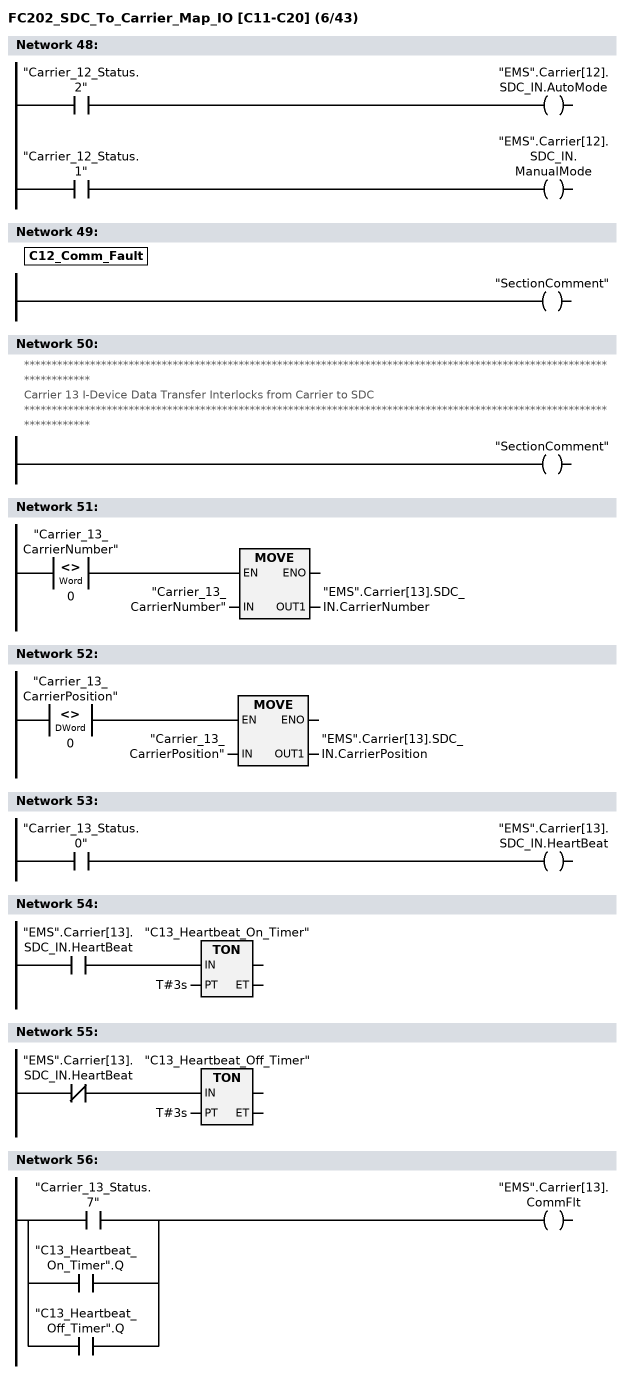
   RUNG wire#powerrail
      Contact( "Carrier_12_Status.2" )
      Coil( "EMS".Carrier[12].SDC_IN.AutoMode )
   END_RUNG
   RUNG wire#powerrail
      Contact( "Carrier_12_Status.1" )
      Coil( "EMS".Carrier[12].SDC_IN.ManualMode )
   END_RUNG
   // the same network as SCL:
   "EMS".Carrier[12].SDC_IN.AutoMode := "Carrier_12_Status.2";
   "EMS".Carrier[12].SDC_IN.ManualMode := "Carrier_12_Status.1";
END_REGION

REGION Network 49
   Label( C12_Comm_Fault )
   RUNG wire#powerrail
      Coil( "SectionComment" )
   END_RUNG
   // the same network as SCL:
   C12_Comm_Fault:
   "SectionComment" := TRUE;
END_REGION

REGION Network 50
   // **********************************************************************************************************************
   // 
   // Carrier 13 I-Device Data Transfer Interlocks from Carrier to SDC
   // 
   // **********************************************************************************************************************
   RUNG wire#powerrail
      Coil( "SectionComment" )
   END_RUNG
   // the same network as SCL:
   "SectionComment" := TRUE;
END_REGION

REGION Network 51
   RUNG wire#powerrail
      { S7_Templates := "SrcType := Word" } NE_Contact(in1 := "Carrier_13_CarrierNumber", in2 := 0)
      Move(in := "Carrier_13_CarrierNumber", out1 => "EMS".Carrier[13].SDC_IN.CarrierNumber)
   END_RUNG
   // the same network as SCL:
   IF "Carrier_13_CarrierNumber" <> 0 THEN
       "EMS".Carrier[13].SDC_IN.CarrierNumber := "Carrier_13_CarrierNumber";
   END_IF;
END_REGION

REGION Network 52
   RUNG wire#powerrail
      { S7_Templates := "SrcType := DWord" } NE_Contact(in1 := "Carrier_13_CarrierPosition", in2 := 0)
      Move(in := "Carrier_13_CarrierPosition", out1 => "EMS".Carrier[13].SDC_IN.CarrierPosition)
   END_RUNG
   // the same network as SCL:
   IF "Carrier_13_CarrierPosition" <> 0 THEN
       "EMS".Carrier[13].SDC_IN.CarrierPosition := "Carrier_13_CarrierPosition";
   END_IF;
END_REGION

REGION Network 53
   RUNG wire#powerrail
      Contact( "Carrier_13_Status.0" )
      Coil( "EMS".Carrier[13].SDC_IN.HeartBeat )
   END_RUNG
   // the same network as SCL:
   "EMS".Carrier[13].SDC_IN.HeartBeat := "Carrier_13_Status.0";
END_REGION

REGION Network 54
   "C13_Heartbeat_On_Timer".TON(IN := "EMS".Carrier[13].SDC_IN.HeartBeat, PT := T#3s);
END_REGION

REGION Network 55
   "C13_Heartbeat_Off_Timer".TON(IN := NOT "EMS".Carrier[13].SDC_IN.HeartBeat, PT := T#3s);
END_REGION

REGION Network 56
   RUNG wire#powerrail
      Contact( "Carrier_13_Status.7" )
      wire#w1
      Coil( "EMS".Carrier[13].CommFlt )
   END_RUNG
   RUNG wire#powerrail
      Contact( "C13_Heartbeat_On_Timer".Q )
   END_RUNG wire#w1
   RUNG wire#powerrail
      Contact( "C13_Heartbeat_Off_Timer".Q )
   END_RUNG wire#w1
   // the same network as SCL:
   "EMS".Carrier[13].CommFlt := "Carrier_13_Status.7" OR "C13_Heartbeat_On_Timer".Q OR "C13_Heartbeat_Off_Timer".Q;
END_REGION

REGION Network 57
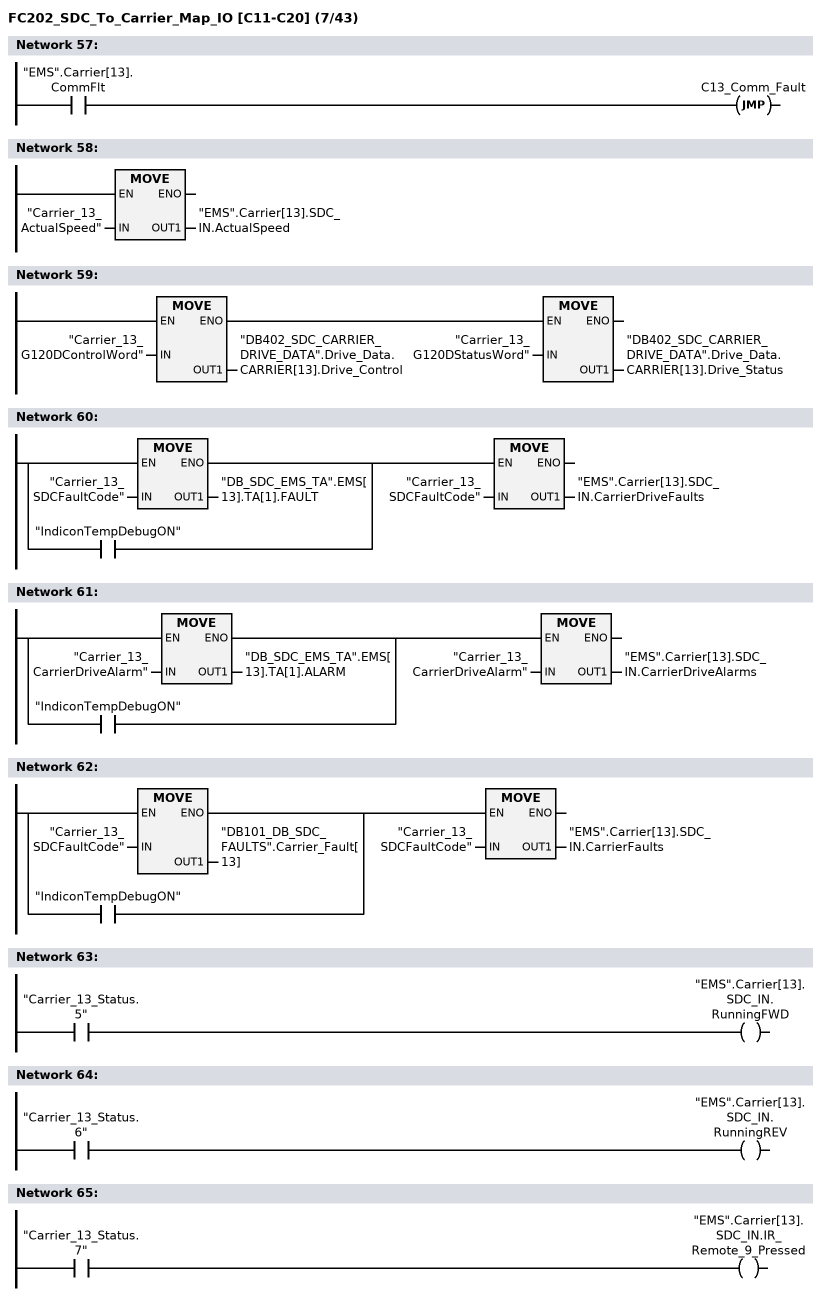
   RUNG wire#powerrail
      Contact( "EMS".Carrier[13].CommFlt )
      JumpCoil( C13_Comm_Fault )
   END_RUNG
   // the same network as SCL:
   IF "EMS".Carrier[13].CommFlt THEN GOTO C13_Comm_Fault; END_IF;
END_REGION

REGION Network 58
   RUNG wire#powerrail
      Move(in := "Carrier_13_ActualSpeed", out1 => "EMS".Carrier[13].SDC_IN.ActualSpeed)
   END_RUNG
   // the same network as SCL:
   "EMS".Carrier[13].SDC_IN.ActualSpeed := "Carrier_13_ActualSpeed";
END_REGION

REGION Network 59
   RUNG wire#powerrail
      Move(in := "Carrier_13_G120DControlWord", out1 => "DB402_SDC_CARRIER_DRIVE_DATA".Drive_Data.CARRIER[13].Drive_Control)
      Move(in := "Carrier_13_G120DStatusWord", out1 => "DB402_SDC_CARRIER_DRIVE_DATA".Drive_Data.CARRIER[13].Drive_Status)
   END_RUNG
   // the same network as SCL:
   "DB402_SDC_CARRIER_DRIVE_DATA".Drive_Data.CARRIER[13].Drive_Control := "Carrier_13_G120DControlWord";
   "DB402_SDC_CARRIER_DRIVE_DATA".Drive_Data.CARRIER[13].Drive_Status := "Carrier_13_G120DStatusWord";
END_REGION

REGION Network 60
   RUNG wire#powerrail
      Move(in := "Carrier_13_SDCFaultCode", out1 => "DB_SDC_EMS_TA".EMS[13].TA[1].FAULT)
      wire#w1
      Move(in := "Carrier_13_SDCFaultCode", out1 => "EMS".Carrier[13].SDC_IN.CarrierDriveFaults)
   END_RUNG
   RUNG wire#powerrail
      Contact( "IndiconTempDebugON" )
   END_RUNG wire#w1
   // the same network as SCL:
   "DB_SDC_EMS_TA".EMS[13].TA[1].FAULT := "Carrier_13_SDCFaultCode";
   IF TRUE OR "IndiconTempDebugON" THEN
       "EMS".Carrier[13].SDC_IN.CarrierDriveFaults := "Carrier_13_SDCFaultCode";
   END_IF;
END_REGION

REGION Network 61
   RUNG wire#powerrail
      Move(in := "Carrier_13_CarrierDriveAlarm", out1 => "DB_SDC_EMS_TA".EMS[13].TA[1].ALARM)
      wire#w1
      Move(in := "Carrier_13_CarrierDriveAlarm", out1 => "EMS".Carrier[13].SDC_IN.CarrierDriveAlarms)
   END_RUNG
   RUNG wire#powerrail
      Contact( "IndiconTempDebugON" )
   END_RUNG wire#w1
   // the same network as SCL:
   "DB_SDC_EMS_TA".EMS[13].TA[1].ALARM := "Carrier_13_CarrierDriveAlarm";
   IF TRUE OR "IndiconTempDebugON" THEN
       "EMS".Carrier[13].SDC_IN.CarrierDriveAlarms := "Carrier_13_CarrierDriveAlarm";
   END_IF;
END_REGION

REGION Network 62
   RUNG wire#powerrail
      Move(in := "Carrier_13_SDCFaultCode", out1 => "DB101_DB_SDC_FAULTS".Carrier_Fault[13])
      wire#w1
      Move(in := "Carrier_13_SDCFaultCode", out1 => "EMS".Carrier[13].SDC_IN.CarrierFaults)
   END_RUNG
   RUNG wire#powerrail
      Contact( "IndiconTempDebugON" )
   END_RUNG wire#w1
   // the same network as SCL:
   "DB101_DB_SDC_FAULTS".Carrier_Fault[13] := "Carrier_13_SDCFaultCode";
   IF TRUE OR "IndiconTempDebugON" THEN
       "EMS".Carrier[13].SDC_IN.CarrierFaults := "Carrier_13_SDCFaultCode";
   END_IF;
END_REGION

REGION Network 63
   RUNG wire#powerrail
      Contact( "Carrier_13_Status.5" )
      Coil( "EMS".Carrier[13].SDC_IN.RunningFWD )
   END_RUNG
   // the same network as SCL:
   "EMS".Carrier[13].SDC_IN.RunningFWD := "Carrier_13_Status.5";
END_REGION

REGION Network 64
   RUNG wire#powerrail
      Contact( "Carrier_13_Status.6" )
      Coil( "EMS".Carrier[13].SDC_IN.RunningREV )
   END_RUNG
   // the same network as SCL:
   "EMS".Carrier[13].SDC_IN.RunningREV := "Carrier_13_Status.6";
END_REGION

REGION Network 65
   RUNG wire#powerrail
      Contact( "Carrier_13_Status.7" )
      Coil( "EMS".Carrier[13].SDC_IN.IR_Remote_9_Pressed )
   END_RUNG
   // the same network as SCL:
   "EMS".Carrier[13].SDC_IN.IR_Remote_9_Pressed := "Carrier_13_Status.7";
END_REGION

REGION Network 66
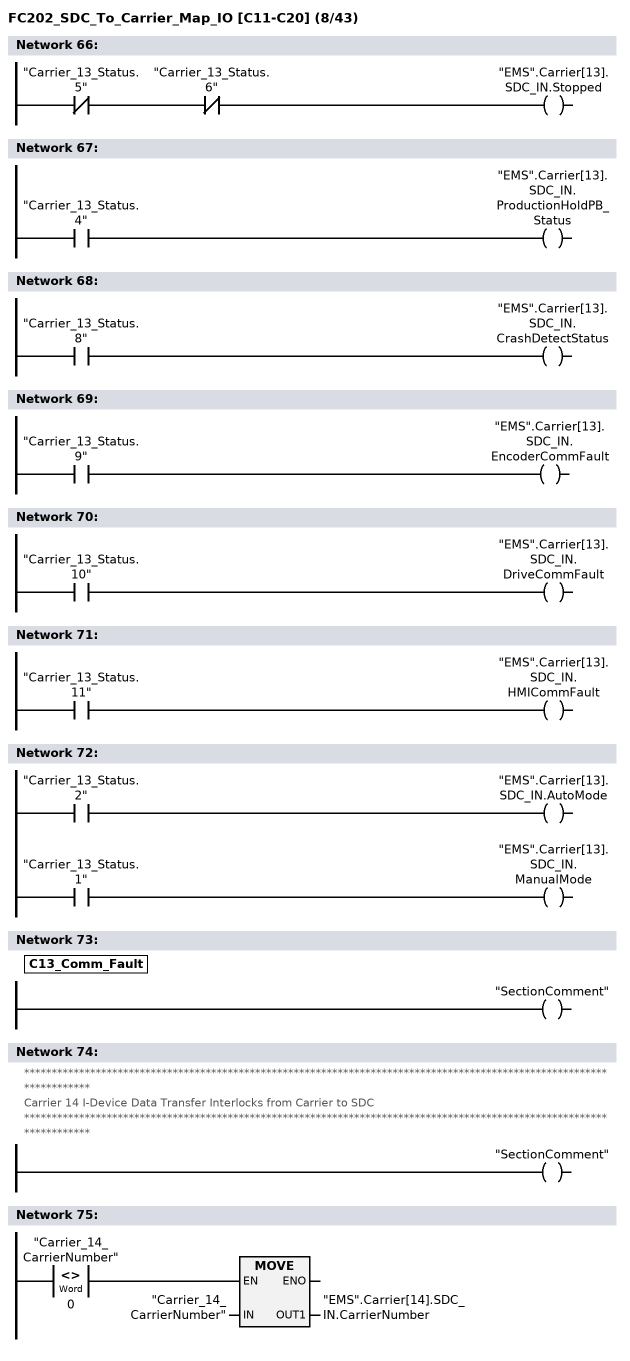
   RUNG wire#powerrail
      I_Contact( "Carrier_13_Status.5" )
      I_Contact( "Carrier_13_Status.6" )
      Coil( "EMS".Carrier[13].SDC_IN.Stopped )
   END_RUNG
   // the same network as SCL:
   "EMS".Carrier[13].SDC_IN.Stopped := NOT "Carrier_13_Status.5" AND NOT "Carrier_13_Status.6";
END_REGION

REGION Network 67
   RUNG wire#powerrail
      Contact( "Carrier_13_Status.4" )
      Coil( "EMS".Carrier[13].SDC_IN.ProductionHoldPB_Status )
   END_RUNG
   // the same network as SCL:
   "EMS".Carrier[13].SDC_IN.ProductionHoldPB_Status := "Carrier_13_Status.4";
END_REGION

REGION Network 68
   RUNG wire#powerrail
      Contact( "Carrier_13_Status.8" )
      Coil( "EMS".Carrier[13].SDC_IN.CrashDetectStatus )
   END_RUNG
   // the same network as SCL:
   "EMS".Carrier[13].SDC_IN.CrashDetectStatus := "Carrier_13_Status.8";
END_REGION

REGION Network 69
   RUNG wire#powerrail
      Contact( "Carrier_13_Status.9" )
      Coil( "EMS".Carrier[13].SDC_IN.EncoderCommFault )
   END_RUNG
   // the same network as SCL:
   "EMS".Carrier[13].SDC_IN.EncoderCommFault := "Carrier_13_Status.9";
END_REGION

REGION Network 70
   RUNG wire#powerrail
      Contact( "Carrier_13_Status.10" )
      Coil( "EMS".Carrier[13].SDC_IN.DriveCommFault )
   END_RUNG
   // the same network as SCL:
   "EMS".Carrier[13].SDC_IN.DriveCommFault := "Carrier_13_Status.10";
END_REGION

REGION Network 71
   RUNG wire#powerrail
      Contact( "Carrier_13_Status.11" )
      Coil( "EMS".Carrier[13].SDC_IN.HMICommFault )
   END_RUNG
   // the same network as SCL:
   "EMS".Carrier[13].SDC_IN.HMICommFault := "Carrier_13_Status.11";
END_REGION

REGION Network 72
   RUNG wire#powerrail
      Contact( "Carrier_13_Status.2" )
      Coil( "EMS".Carrier[13].SDC_IN.AutoMode )
   END_RUNG
   RUNG wire#powerrail
      Contact( "Carrier_13_Status.1" )
      Coil( "EMS".Carrier[13].SDC_IN.ManualMode )
   END_RUNG
   // the same network as SCL:
   "EMS".Carrier[13].SDC_IN.AutoMode := "Carrier_13_Status.2";
   "EMS".Carrier[13].SDC_IN.ManualMode := "Carrier_13_Status.1";
END_REGION

REGION Network 73
   Label( C13_Comm_Fault )
   RUNG wire#powerrail
      Coil( "SectionComment" )
   END_RUNG
   // the same network as SCL:
   C13_Comm_Fault:
   "SectionComment" := TRUE;
END_REGION

REGION Network 74
   // **********************************************************************************************************************
   // 
   // Carrier 14 I-Device Data Transfer Interlocks from Carrier to SDC
   // 
   // **********************************************************************************************************************
   RUNG wire#powerrail
      Coil( "SectionComment" )
   END_RUNG
   // the same network as SCL:
   "SectionComment" := TRUE;
END_REGION

REGION Network 75
   RUNG wire#powerrail
      { S7_Templates := "SrcType := Word" } NE_Contact(in1 := "Carrier_14_CarrierNumber", in2 := 0)
      Move(in := "Carrier_14_CarrierNumber", out1 => "EMS".Carrier[14].SDC_IN.CarrierNumber)
   END_RUNG
   // the same network as SCL:
   IF "Carrier_14_CarrierNumber" <> 0 THEN
       "EMS".Carrier[14].SDC_IN.CarrierNumber := "Carrier_14_CarrierNumber";
   END_IF;
END_REGION

REGION Network 76
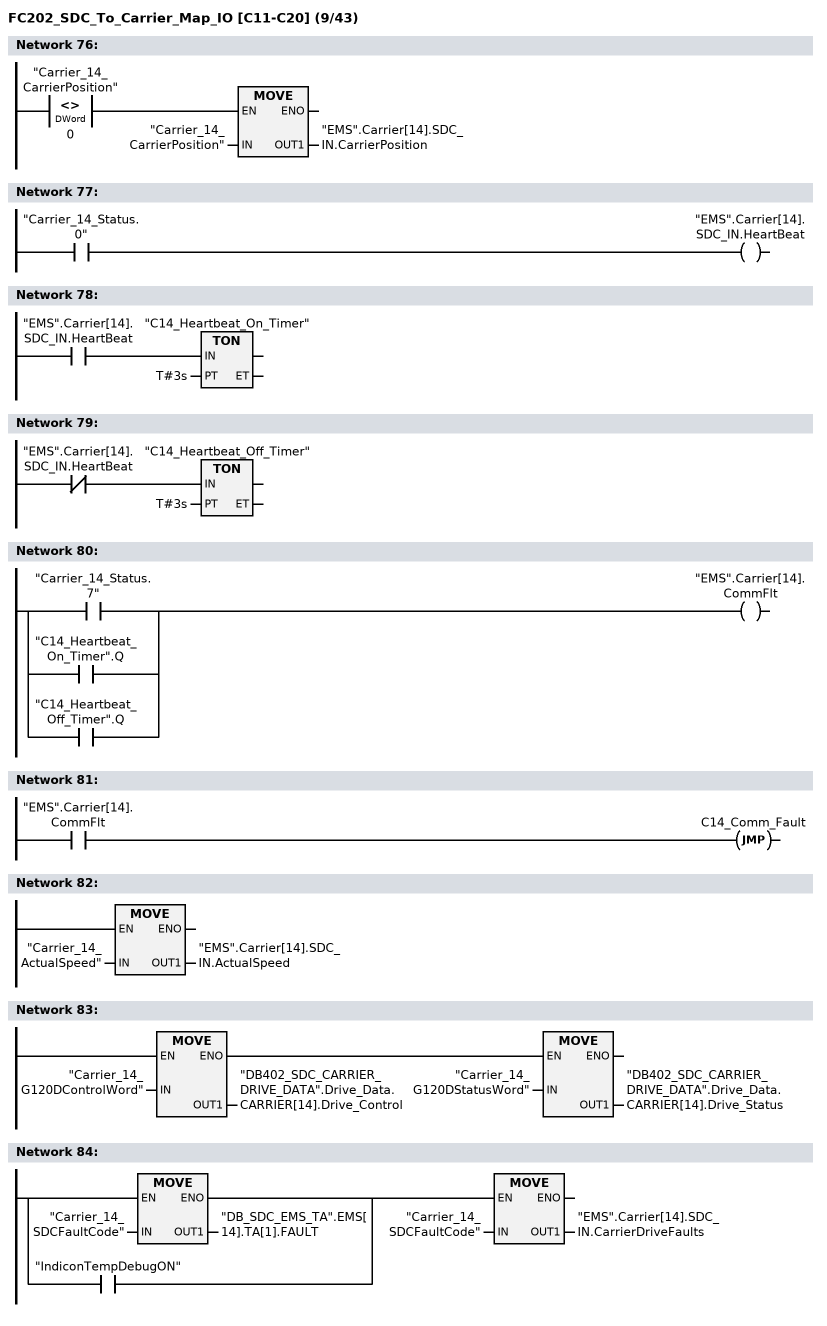
   RUNG wire#powerrail
      { S7_Templates := "SrcType := DWord" } NE_Contact(in1 := "Carrier_14_CarrierPosition", in2 := 0)
      Move(in := "Carrier_14_CarrierPosition", out1 => "EMS".Carrier[14].SDC_IN.CarrierPosition)
   END_RUNG
   // the same network as SCL:
   IF "Carrier_14_CarrierPosition" <> 0 THEN
       "EMS".Carrier[14].SDC_IN.CarrierPosition := "Carrier_14_CarrierPosition";
   END_IF;
END_REGION

REGION Network 77
   RUNG wire#powerrail
      Contact( "Carrier_14_Status.0" )
      Coil( "EMS".Carrier[14].SDC_IN.HeartBeat )
   END_RUNG
   // the same network as SCL:
   "EMS".Carrier[14].SDC_IN.HeartBeat := "Carrier_14_Status.0";
END_REGION

REGION Network 78
   "C14_Heartbeat_On_Timer".TON(IN := "EMS".Carrier[14].SDC_IN.HeartBeat, PT := T#3s);
END_REGION

REGION Network 79
   "C14_Heartbeat_Off_Timer".TON(IN := NOT "EMS".Carrier[14].SDC_IN.HeartBeat, PT := T#3s);
END_REGION

REGION Network 80
   RUNG wire#powerrail
      Contact( "Carrier_14_Status.7" )
      wire#w1
      Coil( "EMS".Carrier[14].CommFlt )
   END_RUNG
   RUNG wire#powerrail
      Contact( "C14_Heartbeat_On_Timer".Q )
   END_RUNG wire#w1
   RUNG wire#powerrail
      Contact( "C14_Heartbeat_Off_Timer".Q )
   END_RUNG wire#w1
   // the same network as SCL:
   "EMS".Carrier[14].CommFlt := "Carrier_14_Status.7" OR "C14_Heartbeat_On_Timer".Q OR "C14_Heartbeat_Off_Timer".Q;
END_REGION

REGION Network 81
   RUNG wire#powerrail
      Contact( "EMS".Carrier[14].CommFlt )
      JumpCoil( C14_Comm_Fault )
   END_RUNG
   // the same network as SCL:
   IF "EMS".Carrier[14].CommFlt THEN GOTO C14_Comm_Fault; END_IF;
END_REGION

REGION Network 82
   RUNG wire#powerrail
      Move(in := "Carrier_14_ActualSpeed", out1 => "EMS".Carrier[14].SDC_IN.ActualSpeed)
   END_RUNG
   // the same network as SCL:
   "EMS".Carrier[14].SDC_IN.ActualSpeed := "Carrier_14_ActualSpeed";
END_REGION

REGION Network 83
   RUNG wire#powerrail
      Move(in := "Carrier_14_G120DControlWord", out1 => "DB402_SDC_CARRIER_DRIVE_DATA".Drive_Data.CARRIER[14].Drive_Control)
      Move(in := "Carrier_14_G120DStatusWord", out1 => "DB402_SDC_CARRIER_DRIVE_DATA".Drive_Data.CARRIER[14].Drive_Status)
   END_RUNG
   // the same network as SCL:
   "DB402_SDC_CARRIER_DRIVE_DATA".Drive_Data.CARRIER[14].Drive_Control := "Carrier_14_G120DControlWord";
   "DB402_SDC_CARRIER_DRIVE_DATA".Drive_Data.CARRIER[14].Drive_Status := "Carrier_14_G120DStatusWord";
END_REGION

REGION Network 84
   RUNG wire#powerrail
      Move(in := "Carrier_14_SDCFaultCode", out1 => "DB_SDC_EMS_TA".EMS[14].TA[1].FAULT)
      wire#w1
      Move(in := "Carrier_14_SDCFaultCode", out1 => "EMS".Carrier[14].SDC_IN.CarrierDriveFaults)
   END_RUNG
   RUNG wire#powerrail
      Contact( "IndiconTempDebugON" )
   END_RUNG wire#w1
   // the same network as SCL:
   "DB_SDC_EMS_TA".EMS[14].TA[1].FAULT := "Carrier_14_SDCFaultCode";
   IF TRUE OR "IndiconTempDebugON" THEN
       "EMS".Carrier[14].SDC_IN.CarrierDriveFaults := "Carrier_14_SDCFaultCode";
   END_IF;
END_REGION

REGION Network 85
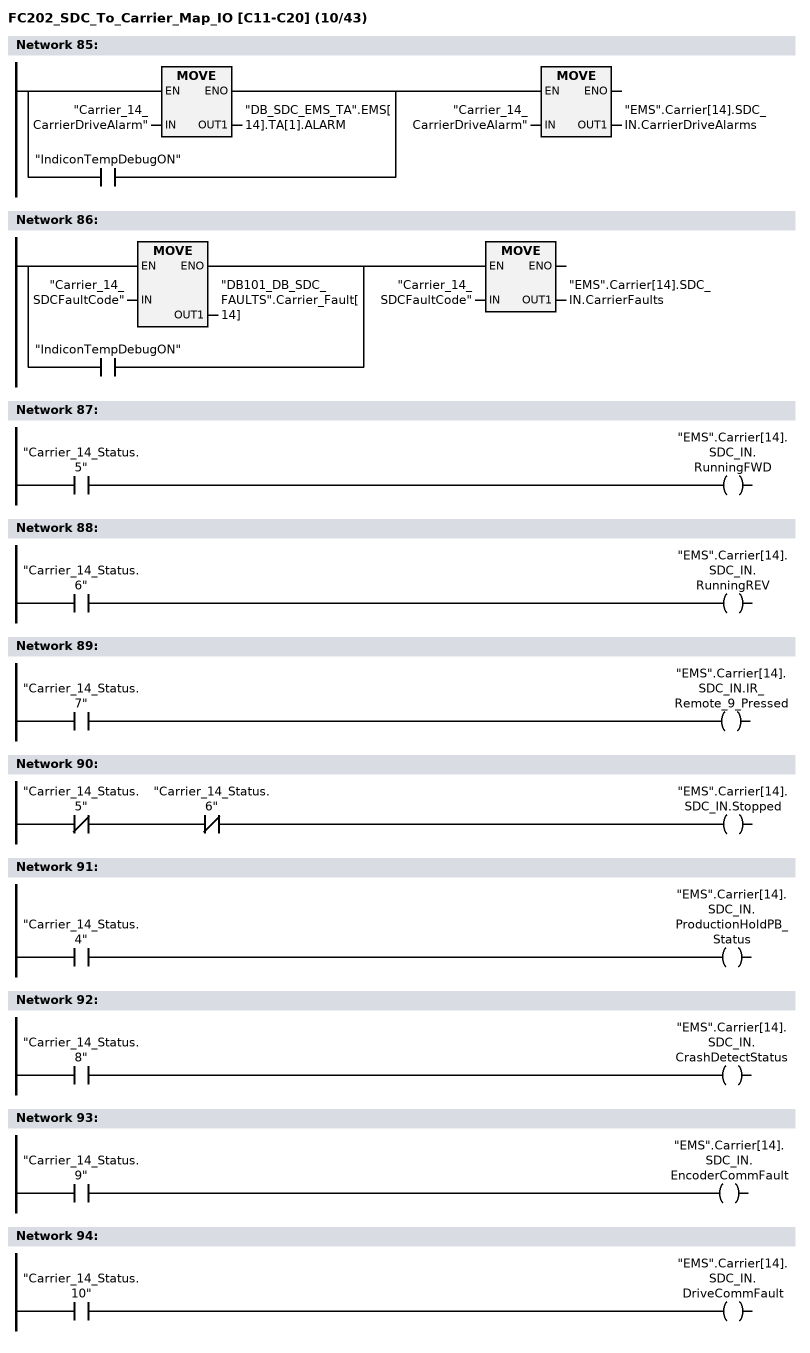
   RUNG wire#powerrail
      Move(in := "Carrier_14_CarrierDriveAlarm", out1 => "DB_SDC_EMS_TA".EMS[14].TA[1].ALARM)
      wire#w1
      Move(in := "Carrier_14_CarrierDriveAlarm", out1 => "EMS".Carrier[14].SDC_IN.CarrierDriveAlarms)
   END_RUNG
   RUNG wire#powerrail
      Contact( "IndiconTempDebugON" )
   END_RUNG wire#w1
   // the same network as SCL:
   "DB_SDC_EMS_TA".EMS[14].TA[1].ALARM := "Carrier_14_CarrierDriveAlarm";
   IF TRUE OR "IndiconTempDebugON" THEN
       "EMS".Carrier[14].SDC_IN.CarrierDriveAlarms := "Carrier_14_CarrierDriveAlarm";
   END_IF;
END_REGION

REGION Network 86
   RUNG wire#powerrail
      Move(in := "Carrier_14_SDCFaultCode", out1 => "DB101_DB_SDC_FAULTS".Carrier_Fault[14])
      wire#w1
      Move(in := "Carrier_14_SDCFaultCode", out1 => "EMS".Carrier[14].SDC_IN.CarrierFaults)
   END_RUNG
   RUNG wire#powerrail
      Contact( "IndiconTempDebugON" )
   END_RUNG wire#w1
   // the same network as SCL:
   "DB101_DB_SDC_FAULTS".Carrier_Fault[14] := "Carrier_14_SDCFaultCode";
   IF TRUE OR "IndiconTempDebugON" THEN
       "EMS".Carrier[14].SDC_IN.CarrierFaults := "Carrier_14_SDCFaultCode";
   END_IF;
END_REGION

REGION Network 87
   RUNG wire#powerrail
      Contact( "Carrier_14_Status.5" )
      Coil( "EMS".Carrier[14].SDC_IN.RunningFWD )
   END_RUNG
   // the same network as SCL:
   "EMS".Carrier[14].SDC_IN.RunningFWD := "Carrier_14_Status.5";
END_REGION

REGION Network 88
   RUNG wire#powerrail
      Contact( "Carrier_14_Status.6" )
      Coil( "EMS".Carrier[14].SDC_IN.RunningREV )
   END_RUNG
   // the same network as SCL:
   "EMS".Carrier[14].SDC_IN.RunningREV := "Carrier_14_Status.6";
END_REGION

REGION Network 89
   RUNG wire#powerrail
      Contact( "Carrier_14_Status.7" )
      Coil( "EMS".Carrier[14].SDC_IN.IR_Remote_9_Pressed )
   END_RUNG
   // the same network as SCL:
   "EMS".Carrier[14].SDC_IN.IR_Remote_9_Pressed := "Carrier_14_Status.7";
END_REGION

REGION Network 90
   RUNG wire#powerrail
      I_Contact( "Carrier_14_Status.5" )
      I_Contact( "Carrier_14_Status.6" )
      Coil( "EMS".Carrier[14].SDC_IN.Stopped )
   END_RUNG
   // the same network as SCL:
   "EMS".Carrier[14].SDC_IN.Stopped := NOT "Carrier_14_Status.5" AND NOT "Carrier_14_Status.6";
END_REGION

REGION Network 91
   RUNG wire#powerrail
      Contact( "Carrier_14_Status.4" )
      Coil( "EMS".Carrier[14].SDC_IN.ProductionHoldPB_Status )
   END_RUNG
   // the same network as SCL:
   "EMS".Carrier[14].SDC_IN.ProductionHoldPB_Status := "Carrier_14_Status.4";
END_REGION

REGION Network 92
   RUNG wire#powerrail
      Contact( "Carrier_14_Status.8" )
      Coil( "EMS".Carrier[14].SDC_IN.CrashDetectStatus )
   END_RUNG
   // the same network as SCL:
   "EMS".Carrier[14].SDC_IN.CrashDetectStatus := "Carrier_14_Status.8";
END_REGION

REGION Network 93
   RUNG wire#powerrail
      Contact( "Carrier_14_Status.9" )
      Coil( "EMS".Carrier[14].SDC_IN.EncoderCommFault )
   END_RUNG
   // the same network as SCL:
   "EMS".Carrier[14].SDC_IN.EncoderCommFault := "Carrier_14_Status.9";
END_REGION

REGION Network 94
   RUNG wire#powerrail
      Contact( "Carrier_14_Status.10" )
      Coil( "EMS".Carrier[14].SDC_IN.DriveCommFault )
   END_RUNG
   // the same network as SCL:
   "EMS".Carrier[14].SDC_IN.DriveCommFault := "Carrier_14_Status.10";
END_REGION

REGION Network 95
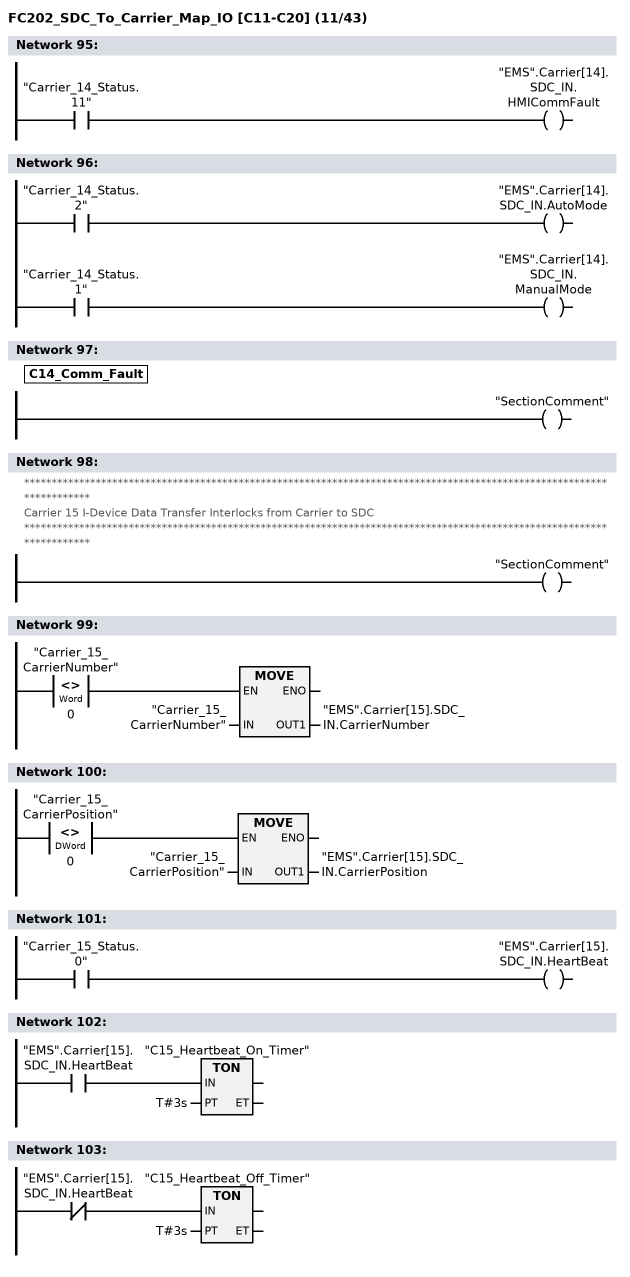
   RUNG wire#powerrail
      Contact( "Carrier_14_Status.11" )
      Coil( "EMS".Carrier[14].SDC_IN.HMICommFault )
   END_RUNG
   // the same network as SCL:
   "EMS".Carrier[14].SDC_IN.HMICommFault := "Carrier_14_Status.11";
END_REGION

REGION Network 96
   RUNG wire#powerrail
      Contact( "Carrier_14_Status.2" )
      Coil( "EMS".Carrier[14].SDC_IN.AutoMode )
   END_RUNG
   RUNG wire#powerrail
      Contact( "Carrier_14_Status.1" )
      Coil( "EMS".Carrier[14].SDC_IN.ManualMode )
   END_RUNG
   // the same network as SCL:
   "EMS".Carrier[14].SDC_IN.AutoMode := "Carrier_14_Status.2";
   "EMS".Carrier[14].SDC_IN.ManualMode := "Carrier_14_Status.1";
END_REGION

REGION Network 97
   Label( C14_Comm_Fault )
   RUNG wire#powerrail
      Coil( "SectionComment" )
   END_RUNG
   // the same network as SCL:
   C14_Comm_Fault:
   "SectionComment" := TRUE;
END_REGION

REGION Network 98
   // **********************************************************************************************************************
   // 
   // Carrier 15 I-Device Data Transfer Interlocks from Carrier to SDC
   // 
   // **********************************************************************************************************************
   RUNG wire#powerrail
      Coil( "SectionComment" )
   END_RUNG
   // the same network as SCL:
   "SectionComment" := TRUE;
END_REGION

REGION Network 99
   RUNG wire#powerrail
      { S7_Templates := "SrcType := Word" } NE_Contact(in1 := "Carrier_15_CarrierNumber", in2 := 0)
      Move(in := "Carrier_15_CarrierNumber", out1 => "EMS".Carrier[15].SDC_IN.CarrierNumber)
   END_RUNG
   // the same network as SCL:
   IF "Carrier_15_CarrierNumber" <> 0 THEN
       "EMS".Carrier[15].SDC_IN.CarrierNumber := "Carrier_15_CarrierNumber";
   END_IF;
END_REGION

REGION Network 100
   RUNG wire#powerrail
      { S7_Templates := "SrcType := DWord" } NE_Contact(in1 := "Carrier_15_CarrierPosition", in2 := 0)
      Move(in := "Carrier_15_CarrierPosition", out1 => "EMS".Carrier[15].SDC_IN.CarrierPosition)
   END_RUNG
   // the same network as SCL:
   IF "Carrier_15_CarrierPosition" <> 0 THEN
       "EMS".Carrier[15].SDC_IN.CarrierPosition := "Carrier_15_CarrierPosition";
   END_IF;
END_REGION

REGION Network 101
   RUNG wire#powerrail
      Contact( "Carrier_15_Status.0" )
      Coil( "EMS".Carrier[15].SDC_IN.HeartBeat )
   END_RUNG
   // the same network as SCL:
   "EMS".Carrier[15].SDC_IN.HeartBeat := "Carrier_15_Status.0";
END_REGION

REGION Network 102
   "C15_Heartbeat_On_Timer".TON(IN := "EMS".Carrier[15].SDC_IN.HeartBeat, PT := T#3s);
END_REGION

REGION Network 103
   "C15_Heartbeat_Off_Timer".TON(IN := NOT "EMS".Carrier[15].SDC_IN.HeartBeat, PT := T#3s);
END_REGION

REGION Network 104
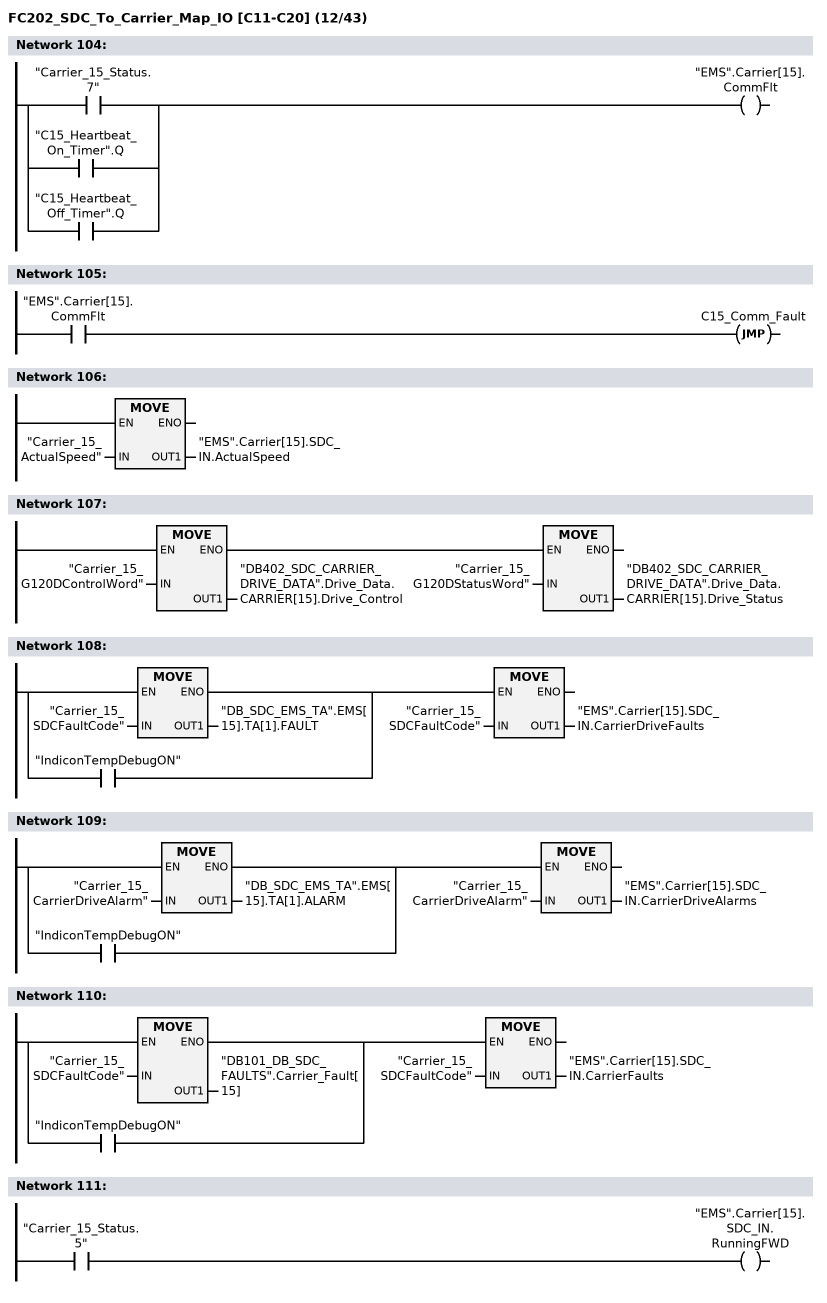
   RUNG wire#powerrail
      Contact( "Carrier_15_Status.7" )
      wire#w1
      Coil( "EMS".Carrier[15].CommFlt )
   END_RUNG
   RUNG wire#powerrail
      Contact( "C15_Heartbeat_On_Timer".Q )
   END_RUNG wire#w1
   RUNG wire#powerrail
      Contact( "C15_Heartbeat_Off_Timer".Q )
   END_RUNG wire#w1
   // the same network as SCL:
   "EMS".Carrier[15].CommFlt := "Carrier_15_Status.7" OR "C15_Heartbeat_On_Timer".Q OR "C15_Heartbeat_Off_Timer".Q;
END_REGION

REGION Network 105
   RUNG wire#powerrail
      Contact( "EMS".Carrier[15].CommFlt )
      JumpCoil( C15_Comm_Fault )
   END_RUNG
   // the same network as SCL:
   IF "EMS".Carrier[15].CommFlt THEN GOTO C15_Comm_Fault; END_IF;
END_REGION

REGION Network 106
   RUNG wire#powerrail
      Move(in := "Carrier_15_ActualSpeed", out1 => "EMS".Carrier[15].SDC_IN.ActualSpeed)
   END_RUNG
   // the same network as SCL:
   "EMS".Carrier[15].SDC_IN.ActualSpeed := "Carrier_15_ActualSpeed";
END_REGION

REGION Network 107
   RUNG wire#powerrail
      Move(in := "Carrier_15_G120DControlWord", out1 => "DB402_SDC_CARRIER_DRIVE_DATA".Drive_Data.CARRIER[15].Drive_Control)
      Move(in := "Carrier_15_G120DStatusWord", out1 => "DB402_SDC_CARRIER_DRIVE_DATA".Drive_Data.CARRIER[15].Drive_Status)
   END_RUNG
   // the same network as SCL:
   "DB402_SDC_CARRIER_DRIVE_DATA".Drive_Data.CARRIER[15].Drive_Control := "Carrier_15_G120DControlWord";
   "DB402_SDC_CARRIER_DRIVE_DATA".Drive_Data.CARRIER[15].Drive_Status := "Carrier_15_G120DStatusWord";
END_REGION

REGION Network 108
   RUNG wire#powerrail
      Move(in := "Carrier_15_SDCFaultCode", out1 => "DB_SDC_EMS_TA".EMS[15].TA[1].FAULT)
      wire#w1
      Move(in := "Carrier_15_SDCFaultCode", out1 => "EMS".Carrier[15].SDC_IN.CarrierDriveFaults)
   END_RUNG
   RUNG wire#powerrail
      Contact( "IndiconTempDebugON" )
   END_RUNG wire#w1
   // the same network as SCL:
   "DB_SDC_EMS_TA".EMS[15].TA[1].FAULT := "Carrier_15_SDCFaultCode";
   IF TRUE OR "IndiconTempDebugON" THEN
       "EMS".Carrier[15].SDC_IN.CarrierDriveFaults := "Carrier_15_SDCFaultCode";
   END_IF;
END_REGION

REGION Network 109
   RUNG wire#powerrail
      Move(in := "Carrier_15_CarrierDriveAlarm", out1 => "DB_SDC_EMS_TA".EMS[15].TA[1].ALARM)
      wire#w1
      Move(in := "Carrier_15_CarrierDriveAlarm", out1 => "EMS".Carrier[15].SDC_IN.CarrierDriveAlarms)
   END_RUNG
   RUNG wire#powerrail
      Contact( "IndiconTempDebugON" )
   END_RUNG wire#w1
   // the same network as SCL:
   "DB_SDC_EMS_TA".EMS[15].TA[1].ALARM := "Carrier_15_CarrierDriveAlarm";
   IF TRUE OR "IndiconTempDebugON" THEN
       "EMS".Carrier[15].SDC_IN.CarrierDriveAlarms := "Carrier_15_CarrierDriveAlarm";
   END_IF;
END_REGION

REGION Network 110
   RUNG wire#powerrail
      Move(in := "Carrier_15_SDCFaultCode", out1 => "DB101_DB_SDC_FAULTS".Carrier_Fault[15])
      wire#w1
      Move(in := "Carrier_15_SDCFaultCode", out1 => "EMS".Carrier[15].SDC_IN.CarrierFaults)
   END_RUNG
   RUNG wire#powerrail
      Contact( "IndiconTempDebugON" )
   END_RUNG wire#w1
   // the same network as SCL:
   "DB101_DB_SDC_FAULTS".Carrier_Fault[15] := "Carrier_15_SDCFaultCode";
   IF TRUE OR "IndiconTempDebugON" THEN
       "EMS".Carrier[15].SDC_IN.CarrierFaults := "Carrier_15_SDCFaultCode";
   END_IF;
END_REGION

REGION Network 111
   RUNG wire#powerrail
      Contact( "Carrier_15_Status.5" )
      Coil( "EMS".Carrier[15].SDC_IN.RunningFWD )
   END_RUNG
   // the same network as SCL:
   "EMS".Carrier[15].SDC_IN.RunningFWD := "Carrier_15_Status.5";
END_REGION

REGION Network 112
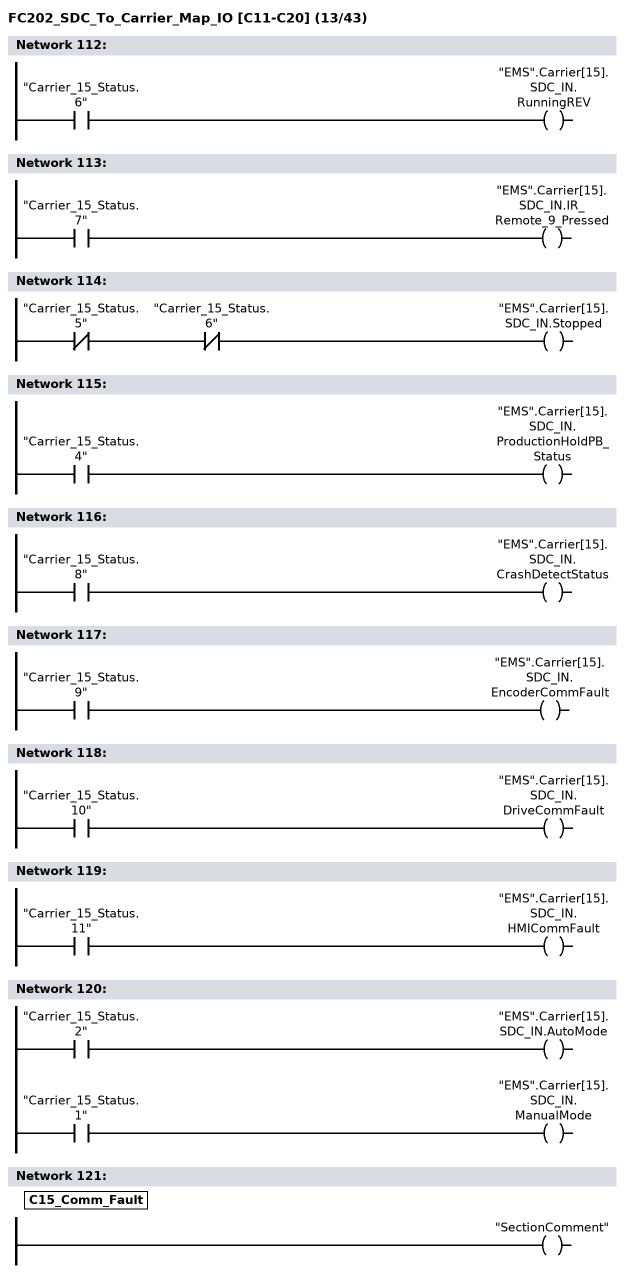
   RUNG wire#powerrail
      Contact( "Carrier_15_Status.6" )
      Coil( "EMS".Carrier[15].SDC_IN.RunningREV )
   END_RUNG
   // the same network as SCL:
   "EMS".Carrier[15].SDC_IN.RunningREV := "Carrier_15_Status.6";
END_REGION

REGION Network 113
   RUNG wire#powerrail
      Contact( "Carrier_15_Status.7" )
      Coil( "EMS".Carrier[15].SDC_IN.IR_Remote_9_Pressed )
   END_RUNG
   // the same network as SCL:
   "EMS".Carrier[15].SDC_IN.IR_Remote_9_Pressed := "Carrier_15_Status.7";
END_REGION

REGION Network 114
   RUNG wire#powerrail
      I_Contact( "Carrier_15_Status.5" )
      I_Contact( "Carrier_15_Status.6" )
      Coil( "EMS".Carrier[15].SDC_IN.Stopped )
   END_RUNG
   // the same network as SCL:
   "EMS".Carrier[15].SDC_IN.Stopped := NOT "Carrier_15_Status.5" AND NOT "Carrier_15_Status.6";
END_REGION

REGION Network 115
   RUNG wire#powerrail
      Contact( "Carrier_15_Status.4" )
      Coil( "EMS".Carrier[15].SDC_IN.ProductionHoldPB_Status )
   END_RUNG
   // the same network as SCL:
   "EMS".Carrier[15].SDC_IN.ProductionHoldPB_Status := "Carrier_15_Status.4";
END_REGION

REGION Network 116
   RUNG wire#powerrail
      Contact( "Carrier_15_Status.8" )
      Coil( "EMS".Carrier[15].SDC_IN.CrashDetectStatus )
   END_RUNG
   // the same network as SCL:
   "EMS".Carrier[15].SDC_IN.CrashDetectStatus := "Carrier_15_Status.8";
END_REGION

REGION Network 117
   RUNG wire#powerrail
      Contact( "Carrier_15_Status.9" )
      Coil( "EMS".Carrier[15].SDC_IN.EncoderCommFault )
   END_RUNG
   // the same network as SCL:
   "EMS".Carrier[15].SDC_IN.EncoderCommFault := "Carrier_15_Status.9";
END_REGION

REGION Network 118
   RUNG wire#powerrail
      Contact( "Carrier_15_Status.10" )
      Coil( "EMS".Carrier[15].SDC_IN.DriveCommFault )
   END_RUNG
   // the same network as SCL:
   "EMS".Carrier[15].SDC_IN.DriveCommFault := "Carrier_15_Status.10";
END_REGION

REGION Network 119
   RUNG wire#powerrail
      Contact( "Carrier_15_Status.11" )
      Coil( "EMS".Carrier[15].SDC_IN.HMICommFault )
   END_RUNG
   // the same network as SCL:
   "EMS".Carrier[15].SDC_IN.HMICommFault := "Carrier_15_Status.11";
END_REGION
